REGION Network 14: Alarm and Warning
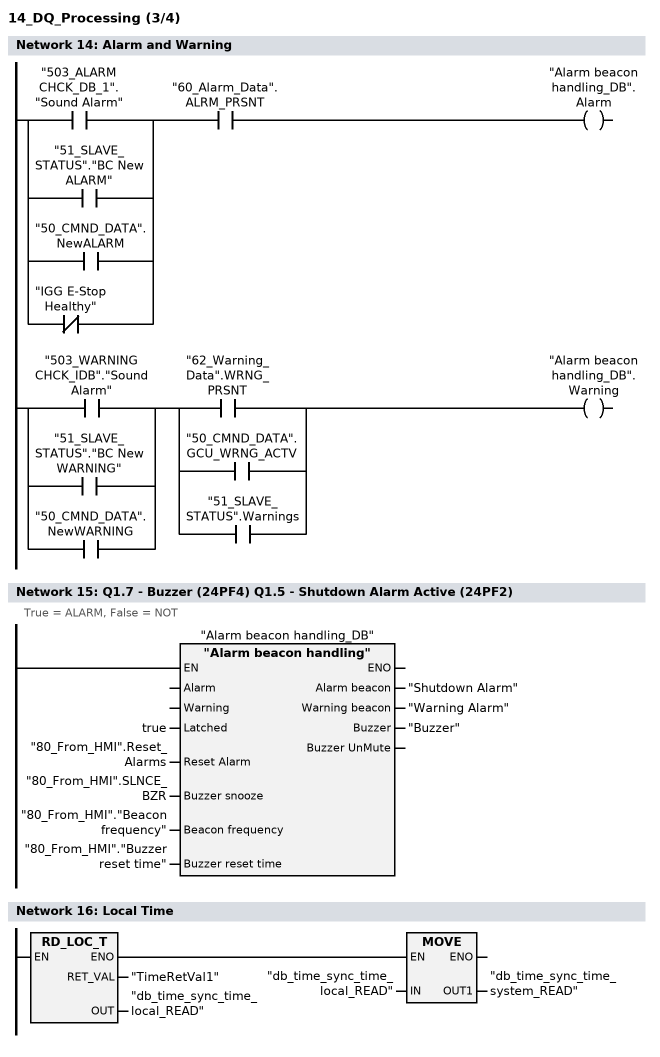
   RUNG wire#powerrail
      Contact( "503_ALARM CHCK_DB_1"."Sound Alarm" )
      wire#w1
      Contact( "60_Alarm_Data".ALRM_PRSNT )
      Coil( "Alarm beacon handling_DB".Alarm )
   END_RUNG
   RUNG wire#powerrail
      Contact( "51_SLAVE_STATUS"."BC New ALARM" )
   END_RUNG wire#w1
   RUNG wire#powerrail
      Contact( "50_CMND_DATA".NewALARM )
   END_RUNG wire#w1
   RUNG wire#powerrail
      I_Contact( "IGG E-Stop Healthy" )
   END_RUNG wire#w1
   RUNG wire#powerrail
      Contact( "503_WARNING CHCK_IDB"."Sound Alarm" )
      wire#w2
      Contact( "62_Warning_Data".WRNG_PRSNT )
      wire#w3
      Coil( "Alarm beacon handling_DB".Warning )
   END_RUNG
   RUNG wire#powerrail
      Contact( "51_SLAVE_STATUS"."BC New WARNING" )
   END_RUNG wire#w2
   RUNG wire#powerrail
      Contact( "50_CMND_DATA".NewWARNING )
   END_RUNG wire#w2
   RUNG wire#w2
      Contact( "50_CMND_DATA".GCU_WRNG_ACTV )
   END_RUNG wire#w3
   RUNG wire#w2
      Contact( "51_SLAVE_STATUS".Warnings )
   END_RUNG wire#w3
   // the same network as SCL:
   "Alarm beacon handling_DB".Alarm := ("503_ALARM CHCK_DB_1"."Sound Alarm" OR "51_SLAVE_STATUS"."BC New ALARM" OR "50_CMND_DATA".NewALARM OR NOT "IGG E-Stop Healthy") AND "60_Alarm_Data".ALRM_PRSNT;
   "Alarm beacon handling_DB".Warning := ("503_WARNING CHCK_IDB"."Sound Alarm" OR "51_SLAVE_STATUS"."BC New WARNING" OR "50_CMND_DATA".NewWARNING) AND ("62_Warning_Data".WRNG_PRSNT OR "50_CMND_DATA".GCU_WRNG_ACTV OR "51_SLAVE_STATUS".Warnings);
END_REGION

REGION Network 15: Q1.7 - Buzzer (24PF4) Q1.5 - Shutdown Alarm Active (24PF2)
   // True = ALARM, False = NOT
   RUNG wire#powerrail
      "Alarm beacon handling_DB"(Alarm :=, Warning :=, Latched := true, "Reset Alarm" := "80_From_HMI".Reset_Alarms, "Buzzer snooze" := "80_From_HMI".SLNCE_BZR, "Beacon frequency" := "80_From_HMI"."Beacon frequency", "Buzzer reset time" := "80_From_HMI"."Buzzer reset time", "Alarm beacon" => "Shutdown Alarm", "Warning beacon" => "Warning Alarm", Buzzer => "Buzzer", "Buzzer UnMute" =>)
   END_RUNG
   // the same network as SCL:
   "Alarm beacon handling_DB"(Latched := true,   // "Alarm beacon handling"
                           "Reset Alarm" := "80_From_HMI".Reset_Alarms,
                           "Buzzer snooze" := "80_From_HMI".SLNCE_BZR,
                           "Beacon frequency" := "80_From_HMI"."Beacon frequency",
                           "Buzzer reset time" := "80_From_HMI"."Buzzer reset time",
                           "Alarm beacon" => "Shutdown Alarm",
                           "Warning beacon" => "Warning Alarm",
                           Buzzer => "Buzzer");
END_REGION

REGION Network 16: Local Time
   // ENO of a box is taken as its EN; it also drops when the box reports an error
   "TimeRetVal1" := RD_LOC_T(OUT => "db_time_sync_time_local_READ");
   "db_time_sync_time_system_READ" := "db_time_sync_time_local_READ";
END_REGION

REGION Network 17: WRITE LOCAL TIME
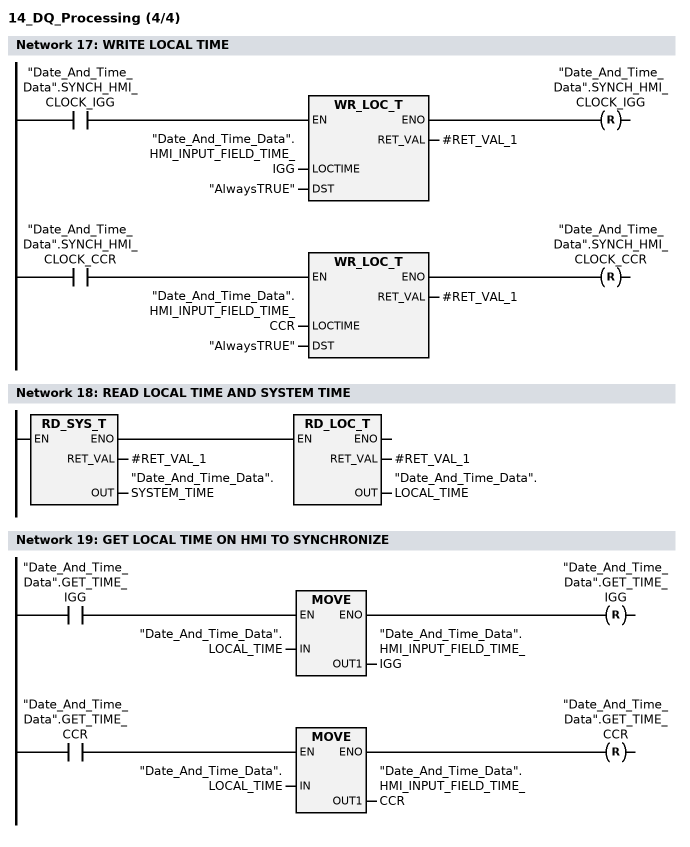
   // ENO of a box is taken as its EN; it also drops when the box reports an error
   #_w1 := "Date_And_Time_Data".SYNCH_HMI_CLOCK_IGG;
   IF #_w1 THEN
       #RET_VAL_1 := WR_LOC_T(LOCTIME := "Date_And_Time_Data".HMI_INPUT_FIELD_TIME_IGG, DST := "AlwaysTRUE");
       "Date_And_Time_Data".SYNCH_HMI_CLOCK_IGG := FALSE;
   END_IF;
   #_w2 := "Date_And_Time_Data".SYNCH_HMI_CLOCK_CCR;
   IF #_w2 THEN
       #RET_VAL_1 := WR_LOC_T(LOCTIME := "Date_And_Time_Data".HMI_INPUT_FIELD_TIME_CCR, DST := "AlwaysTRUE");
       "Date_And_Time_Data".SYNCH_HMI_CLOCK_CCR := FALSE;
   END_IF;
END_REGION

REGION Network 18: READ LOCAL TIME AND SYSTEM TIME
   // ENO of a box is taken as its EN; it also drops when the box reports an error
   #RET_VAL_1 := RD_SYS_T(OUT => "Date_And_Time_Data".SYSTEM_TIME);
   #RET_VAL_1 := RD_LOC_T(OUT => "Date_And_Time_Data".LOCAL_TIME);
END_REGION

REGION Network 19: GET LOCAL TIME ON HMI TO SYNCHRONIZE
   RUNG wire#powerrail
      Contact( "Date_And_Time_Data".GET_TIME_IGG )
      Move(in := "Date_And_Time_Data".LOCAL_TIME, out1 => "Date_And_Time_Data".HMI_INPUT_FIELD_TIME_IGG)
      R_Coil( "Date_And_Time_Data".GET_TIME_IGG )
   END_RUNG
   RUNG wire#powerrail
      Contact( "Date_And_Time_Data".GET_TIME_CCR )
      Move(in := "Date_And_Time_Data".LOCAL_TIME, out1 => "Date_And_Time_Data".HMI_INPUT_FIELD_TIME_CCR)
      R_Coil( "Date_And_Time_Data".GET_TIME_CCR )
   END_RUNG
   // the same network as SCL:
   IF "Date_And_Time_Data".GET_TIME_IGG THEN
       "Date_And_Time_Data".HMI_INPUT_FIELD_TIME_IGG := "Date_And_Time_Data".LOCAL_TIME;
       "Date_And_Time_Data".GET_TIME_IGG := FALSE;
   END_IF;
   IF "Date_And_Time_Data".GET_TIME_CCR THEN
       "Date_And_Time_Data".HMI_INPUT_FIELD_TIME_CCR := "Date_And_Time_Data".LOCAL_TIME;
       "Date_And_Time_Data".GET_TIME_CCR := FALSE;
   END_IF;
END_REGION
END_FUNCTION

FUNCTION "16_AQ_Processing" : Void   // FC16, LAD
TITLE = Analogue Output Processing
{ S7_Optimized_Access := 'TRUE' }
AUTHOR : JRS
VERSION : 0.1
// To process code outputs prior to physical connection
BEGIN

REGION Network 1: QW98 - Vent Valve Position Control (CV-403)
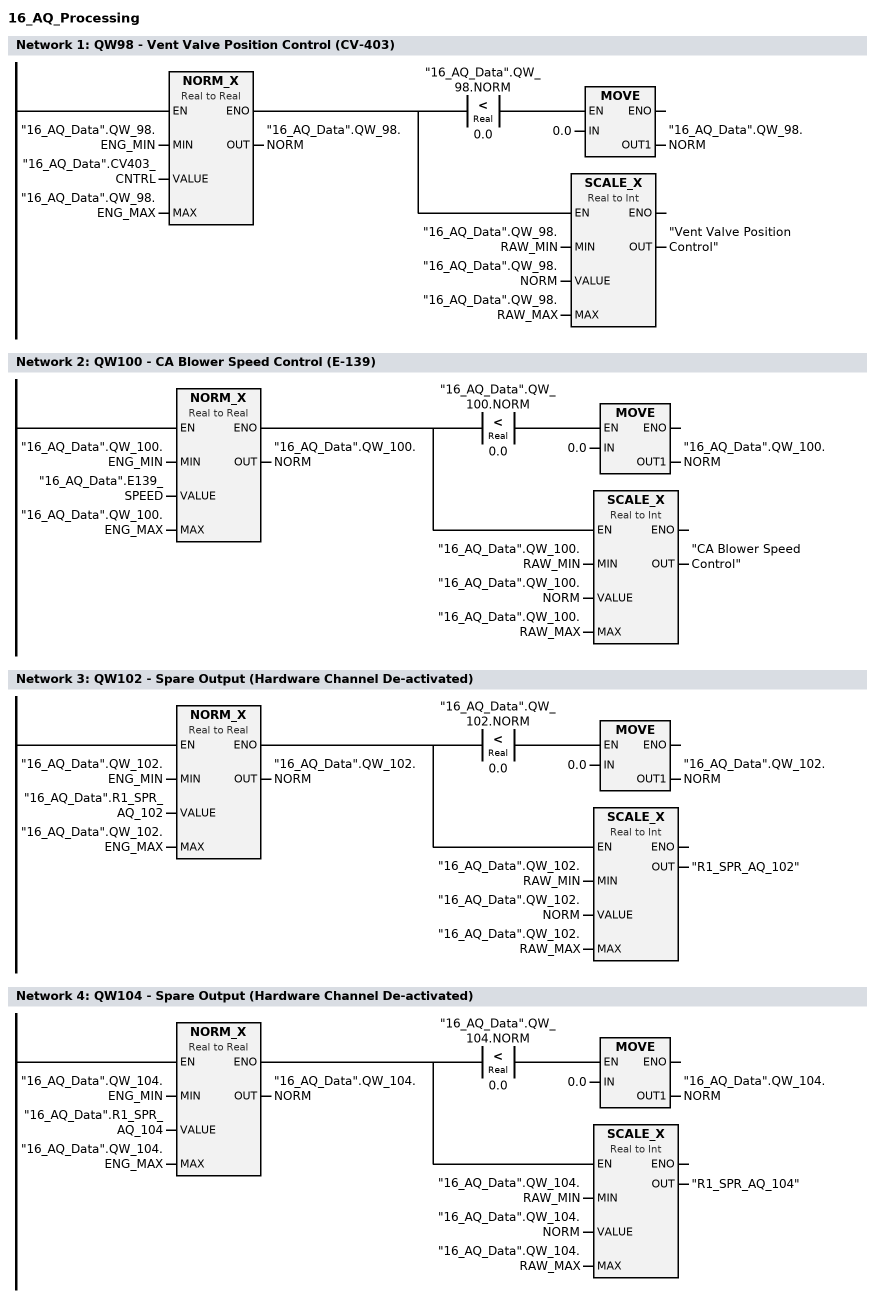
   RUNG wire#powerrail
      { S7_Templates := "[SrcType := Real, DestType := Real]" } Normalize(min := "16_AQ_Data".QW_98.ENG_MIN, value := "16_AQ_Data".CV403_CNTRL, max := "16_AQ_Data".QW_98.ENG_MAX, out => "16_AQ_Data".QW_98.NORM)
      wire#w1
      { S7_Templates := "SrcType := Real" } LT_Contact(in1 := "16_AQ_Data".QW_98.NORM, in2 := 0.0)
      Move(in := 0.0, out1 => "16_AQ_Data".QW_98.NORM)
   END_RUNG
   RUNG wire#w1
      { S7_Templates := "[SrcType := Real, DestType := Int]" } Scale(min := "16_AQ_Data".QW_98.RAW_MIN, value := "16_AQ_Data".QW_98.NORM, max := "16_AQ_Data".QW_98.RAW_MAX, out => "Vent Valve Position Control")
   END_RUNG
   // the same network as SCL:
   "16_AQ_Data".QW_98.NORM := NORM_X(MIN := "16_AQ_Data".QW_98.ENG_MIN, VALUE := "16_AQ_Data".CV403_CNTRL, MAX := "16_AQ_Data".QW_98.ENG_MAX);
   IF "16_AQ_Data".QW_98.NORM < 0.0 THEN "16_AQ_Data".QW_98.NORM := 0.0; END_IF;
   "Vent Valve Position Control" := SCALE_X(MIN := "16_AQ_Data".QW_98.RAW_MIN, VALUE := "16_AQ_Data".QW_98.NORM, MAX := "16_AQ_Data".QW_98.RAW_MAX);
END_REGION

REGION Network 2: QW100 - CA Blower Speed Control (E-139)
   RUNG wire#powerrail
      { S7_Templates := "[SrcType := Real, DestType := Real]" } Normalize(min := "16_AQ_Data".QW_100.ENG_MIN, value := "16_AQ_Data".E139_SPEED, max := "16_AQ_Data".QW_100.ENG_MAX, out => "16_AQ_Data".QW_100.NORM)
      wire#w1
      { S7_Templates := "SrcType := Real" } LT_Contact(in1 := "16_AQ_Data".QW_100.NORM, in2 := 0.0)
      Move(in := 0.0, out1 => "16_AQ_Data".QW_100.NORM)
   END_RUNG
   RUNG wire#w1
      { S7_Templates := "[SrcType := Real, DestType := Int]" } Scale(min := "16_AQ_Data".QW_100.RAW_MIN, value := "16_AQ_Data".QW_100.NORM, max := "16_AQ_Data".QW_100.RAW_MAX, out => "CA Blower Speed Control")
   END_RUNG
   // the same network as SCL:
   "16_AQ_Data".QW_100.NORM := NORM_X(MIN := "16_AQ_Data".QW_100.ENG_MIN, VALUE := "16_AQ_Data".E139_SPEED, MAX := "16_AQ_Data".QW_100.ENG_MAX);
   IF "16_AQ_Data".QW_100.NORM < 0.0 THEN "16_AQ_Data".QW_100.NORM := 0.0; END_IF;
   "CA Blower Speed Control" := SCALE_X(MIN := "16_AQ_Data".QW_100.RAW_MIN, VALUE := "16_AQ_Data".QW_100.NORM, MAX := "16_AQ_Data".QW_100.RAW_MAX);
END_REGION

REGION Network 3: QW102 - Spare Output (Hardware Channel De-activated)
   RUNG wire#powerrail
      { S7_Templates := "[SrcType := Real, DestType := Real]" } Normalize(min := "16_AQ_Data".QW_102.ENG_MIN, value := "16_AQ_Data".R1_SPR_AQ_102, max := "16_AQ_Data".QW_102.ENG_MAX, out => "16_AQ_Data".QW_102.NORM)
      wire#w1
      { S7_Templates := "SrcType := Real" } LT_Contact(in1 := "16_AQ_Data".QW_102.NORM, in2 := 0.0)
      Move(in := 0.0, out1 => "16_AQ_Data".QW_102.NORM)
   END_RUNG
   RUNG wire#w1
      { S7_Templates := "[SrcType := Real, DestType := Int]" } Scale(min := "16_AQ_Data".QW_102.RAW_MIN, value := "16_AQ_Data".QW_102.NORM, max := "16_AQ_Data".QW_102.RAW_MAX, out => "R1_SPR_AQ_102")
   END_RUNG
   // the same network as SCL:
   "16_AQ_Data".QW_102.NORM := NORM_X(MIN := "16_AQ_Data".QW_102.ENG_MIN, VALUE := "16_AQ_Data".R1_SPR_AQ_102, MAX := "16_AQ_Data".QW_102.ENG_MAX);
   IF "16_AQ_Data".QW_102.NORM < 0.0 THEN "16_AQ_Data".QW_102.NORM := 0.0; END_IF;
   "R1_SPR_AQ_102" := SCALE_X(MIN := "16_AQ_Data".QW_102.RAW_MIN, VALUE := "16_AQ_Data".QW_102.NORM, MAX := "16_AQ_Data".QW_102.RAW_MAX);
END_REGION

REGION Network 4: QW104 - Spare Output (Hardware Channel De-activated)
   RUNG wire#powerrail
      { S7_Templates := "[SrcType := Real, DestType := Real]" } Normalize(min := "16_AQ_Data".QW_104.ENG_MIN, value := "16_AQ_Data".R1_SPR_AQ_104, max := "16_AQ_Data".QW_104.ENG_MAX, out => "16_AQ_Data".QW_104.NORM)
      wire#w1
      { S7_Templates := "SrcType := Real" } LT_Contact(in1 := "16_AQ_Data".QW_104.NORM, in2 := 0.0)
      Move(in := 0.0, out1 => "16_AQ_Data".QW_104.NORM)
   END_RUNG
   RUNG wire#w1
      { S7_Templates := "[SrcType := Real, DestType := Int]" } Scale(min := "16_AQ_Data".QW_104.RAW_MIN, value := "16_AQ_Data".QW_104.NORM, max := "16_AQ_Data".QW_104.RAW_MAX, out => "R1_SPR_AQ_104")
   END_RUNG
   // the same network as SCL:
   "16_AQ_Data".QW_104.NORM := NORM_X(MIN := "16_AQ_Data".QW_104.ENG_MIN, VALUE := "16_AQ_Data".R1_SPR_AQ_104, MAX := "16_AQ_Data".QW_104.ENG_MAX);
   IF "16_AQ_Data".QW_104.NORM < 0.0 THEN "16_AQ_Data".QW_104.NORM := 0.0; END_IF;
   "R1_SPR_AQ_104" := SCALE_X(MIN := "16_AQ_Data".QW_104.RAW_MIN, VALUE := "16_AQ_Data".QW_104.NORM, MAX := "16_AQ_Data".QW_104.RAW_MAX);
END_REGION
END_FUNCTION

FUNCTION "19_AUTO_CMNDS" : Void   // FC19, LAD
TITLE = Automatic Output Commands
{ S7_Optimized_Access := 'TRUE' }
AUTHOR : JRS
VERSION : 0.1
// To process automatic output commands prior to output processing
   VAR_TEMP   // added for the SCL form of the ladder/FBD networks
      _w1 : Bool;
      _w2 : Bool;
   END_VAR
BEGIN

REGION Network 1: Fuel Pumps Control
   // Demand from sequence     ...changed from 80 to 140
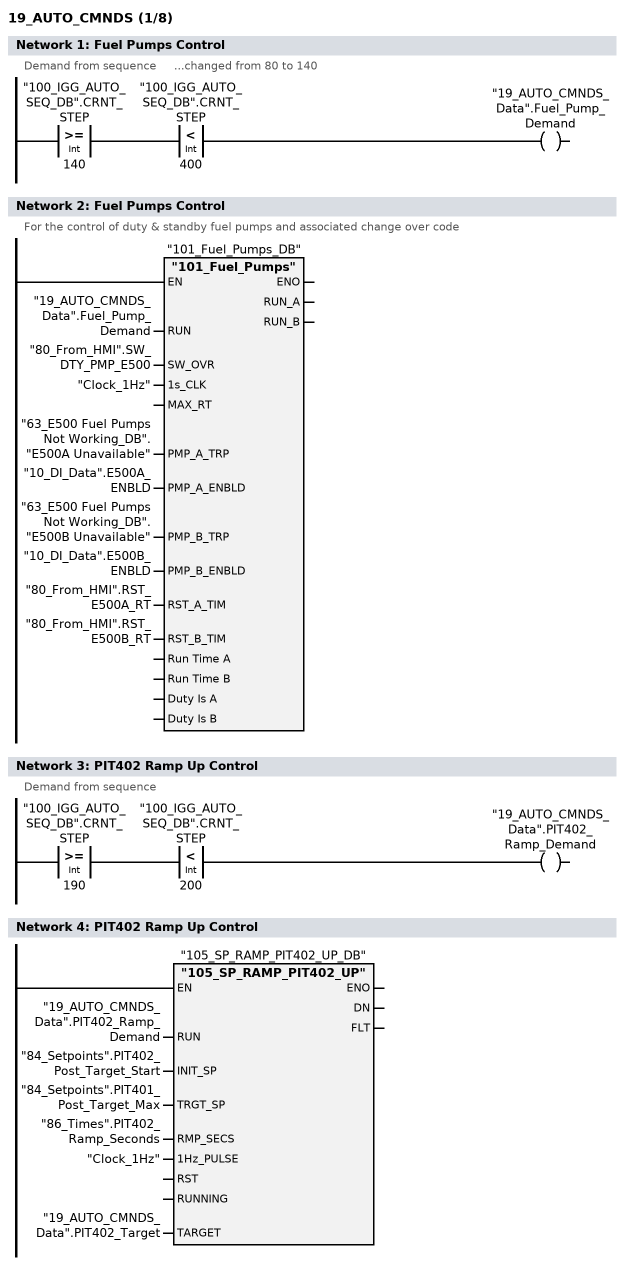
   RUNG wire#powerrail
      { S7_Templates := "SrcType := Int" } GE_Contact(in1 := "100_IGG_AUTO_SEQ_DB".CRNT_STEP, in2 := 140)
      { S7_Templates := "SrcType := Int" } LT_Contact(in1 := "100_IGG_AUTO_SEQ_DB".CRNT_STEP, in2 := 400)
      Coil( "19_AUTO_CMNDS_Data".Fuel_Pump_Demand )
   END_RUNG
   // the same network as SCL:
   "19_AUTO_CMNDS_Data".Fuel_Pump_Demand := ("100_IGG_AUTO_SEQ_DB".CRNT_STEP >= 140) AND ("100_IGG_AUTO_SEQ_DB".CRNT_STEP < 400);
END_REGION

REGION Network 2: Fuel Pumps Control
   // For the control of duty & standby fuel pumps and associated change over code
   RUNG wire#powerrail
      "101_Fuel_Pumps_DB"(RUN := "19_AUTO_CMNDS_Data".Fuel_Pump_Demand, SW_OVR := "80_From_HMI".SW_DTY_PMP_E500, "1s_CLK" := "Clock_1Hz", MAX_RT :=, PMP_A_TRP := "63_E500 Fuel Pumps Not Working_DB"."E500A Unavailable", PMP_A_ENBLD := "10_DI_Data".E500A_ENBLD, PMP_B_TRP := "63_E500 Fuel Pumps Not Working_DB"."E500B Unavailable", PMP_B_ENBLD := "10_DI_Data".E500B_ENBLD, RST_A_TIM := "80_From_HMI".RST_E500A_RT, RST_B_TIM := "80_From_HMI".RST_E500B_RT, "Run Time A" :=, "Run Time B" :=, "Duty Is A" :=, "Duty Is B" :=, RUN_A =>, RUN_B =>)
   END_RUNG
   // the same network as SCL:
   "101_Fuel_Pumps_DB"(RUN := "19_AUTO_CMNDS_Data".Fuel_Pump_Demand,   // "101_Fuel_Pumps"
                       SW_OVR := "80_From_HMI".SW_DTY_PMP_E500,
                       "1s_CLK" := "Clock_1Hz",
                       PMP_A_TRP := "63_E500 Fuel Pumps Not Working_DB"."E500A Unavailable",
                       PMP_A_ENBLD := "10_DI_Data".E500A_ENBLD,
                       PMP_B_TRP := "63_E500 Fuel Pumps Not Working_DB"."E500B Unavailable",
                       PMP_B_ENBLD := "10_DI_Data".E500B_ENBLD,
                       RST_A_TIM := "80_From_HMI".RST_E500A_RT,
                       RST_B_TIM := "80_From_HMI".RST_E500B_RT);
END_REGION

REGION Network 3: PIT402 Ramp Up Control
   // Demand from sequence
   RUNG wire#powerrail
      { S7_Templates := "SrcType := Int" } GE_Contact(in1 := "100_IGG_AUTO_SEQ_DB".CRNT_STEP, in2 := 190)
      { S7_Templates := "SrcType := Int" } LT_Contact(in1 := "100_IGG_AUTO_SEQ_DB".CRNT_STEP, in2 := 200)
      Coil( "19_AUTO_CMNDS_Data".PIT402_Ramp_Demand )
   END_RUNG
   // the same network as SCL:
   "19_AUTO_CMNDS_Data".PIT402_Ramp_Demand := ("100_IGG_AUTO_SEQ_DB".CRNT_STEP >= 190) AND ("100_IGG_AUTO_SEQ_DB".CRNT_STEP < 200);
END_REGION

REGION Network 4: PIT402 Ramp Up Control
   RUNG wire#powerrail
      "105_SP_RAMP_PIT402_UP_DB"(RUN := "19_AUTO_CMNDS_Data".PIT402_Ramp_Demand, INIT_SP := "84_Setpoints".PIT402_Post_Target_Start, TRGT_SP := "84_Setpoints".PIT401_Post_Target_Max, RMP_SECS := "86_Times".PIT402_Ramp_Seconds, "1Hz_PULSE" := "Clock_1Hz", RST :=, RUNNING :=, TARGET := "19_AUTO_CMNDS_Data".PIT402_Target, DN =>, FLT =>)
   END_RUNG
   // the same network as SCL:
   "105_SP_RAMP_PIT402_UP_DB"(RUN := "19_AUTO_CMNDS_Data".PIT402_Ramp_Demand,   // "105_SP_RAMP_PIT402_UP"
                           INIT_SP := "84_Setpoints".PIT402_Post_Target_Start,
                           TRGT_SP := "84_Setpoints".PIT401_Post_Target_Max,
                           RMP_SECS := "86_Times".PIT402_Ramp_Seconds,
                           "1Hz_PULSE" := "Clock_1Hz",
                           TARGET := "19_AUTO_CMNDS_Data".PIT402_Target);
END_REGION

REGION Network 5: PIT402 Ramp Down Control
   // Demand from sequence
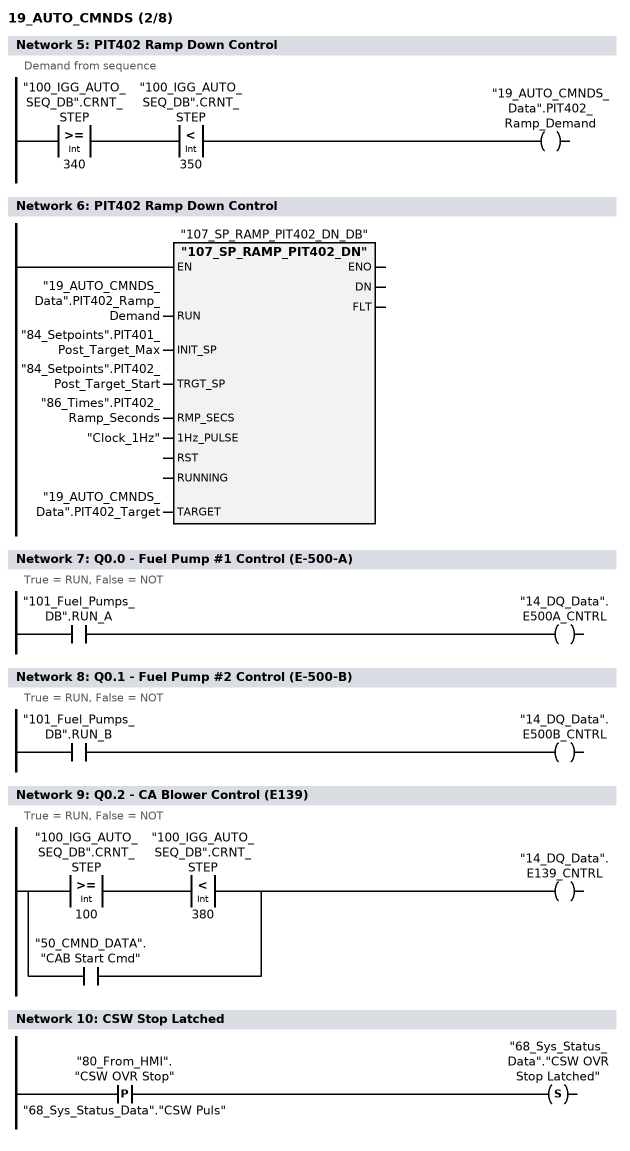
   RUNG wire#powerrail
      { S7_Templates := "SrcType := Int" } GE_Contact(in1 := "100_IGG_AUTO_SEQ_DB".CRNT_STEP, in2 := 340)
      { S7_Templates := "SrcType := Int" } LT_Contact(in1 := "100_IGG_AUTO_SEQ_DB".CRNT_STEP, in2 := 350)
      Coil( "19_AUTO_CMNDS_Data".PIT402_Ramp_Demand )
   END_RUNG
   // the same network as SCL:
   "19_AUTO_CMNDS_Data".PIT402_Ramp_Demand := ("100_IGG_AUTO_SEQ_DB".CRNT_STEP >= 340) AND ("100_IGG_AUTO_SEQ_DB".CRNT_STEP < 350);
END_REGION

REGION Network 6: PIT402 Ramp Down Control
   RUNG wire#powerrail
      "107_SP_RAMP_PIT402_DN_DB"(RUN := "19_AUTO_CMNDS_Data".PIT402_Ramp_Demand, INIT_SP := "84_Setpoints".PIT401_Post_Target_Max, TRGT_SP := "84_Setpoints".PIT402_Post_Target_Start, RMP_SECS := "86_Times".PIT402_Ramp_Seconds, "1Hz_PULSE" := "Clock_1Hz", RST :=, RUNNING :=, TARGET := "19_AUTO_CMNDS_Data".PIT402_Target, DN =>, FLT =>)
   END_RUNG
   // the same network as SCL:
   "107_SP_RAMP_PIT402_DN_DB"(RUN := "19_AUTO_CMNDS_Data".PIT402_Ramp_Demand,   // "107_SP_RAMP_PIT402_DN"
                           INIT_SP := "84_Setpoints".PIT401_Post_Target_Max,
                           TRGT_SP := "84_Setpoints".PIT402_Post_Target_Start,
                           RMP_SECS := "86_Times".PIT402_Ramp_Seconds,
                           "1Hz_PULSE" := "Clock_1Hz",
                           TARGET := "19_AUTO_CMNDS_Data".PIT402_Target);
END_REGION

REGION Network 7: Q0.0 - Fuel Pump #1 Control (E-500-A)
   // True = RUN, False = NOT
   RUNG wire#powerrail
      Contact( "101_Fuel_Pumps_DB".RUN_A )
      Coil( "14_DQ_Data".E500A_CNTRL )
   END_RUNG
   // the same network as SCL:
   "14_DQ_Data".E500A_CNTRL := "101_Fuel_Pumps_DB".RUN_A;
END_REGION

REGION Network 8: Q0.1 - Fuel Pump #2 Control (E-500-B)
   // True = RUN, False = NOT
   RUNG wire#powerrail
      Contact( "101_Fuel_Pumps_DB".RUN_B )
      Coil( "14_DQ_Data".E500B_CNTRL )
   END_RUNG
   // the same network as SCL:
   "14_DQ_Data".E500B_CNTRL := "101_Fuel_Pumps_DB".RUN_B;
END_REGION

REGION Network 9: Q0.2 - CA Blower Control (E139)
   // True = RUN, False = NOT
   RUNG wire#powerrail
      { S7_Templates := "SrcType := Int" } GE_Contact(in1 := "100_IGG_AUTO_SEQ_DB".CRNT_STEP, in2 := 100)
      { S7_Templates := "SrcType := Int" } LT_Contact(in1 := "100_IGG_AUTO_SEQ_DB".CRNT_STEP, in2 := 380)
      wire#w1
      Coil( "14_DQ_Data".E139_CNTRL )
   END_RUNG
   RUNG wire#powerrail
      Contact( "50_CMND_DATA"."CAB Start Cmd" )
   END_RUNG wire#w1
   // the same network as SCL:
   "14_DQ_Data".E139_CNTRL := (("100_IGG_AUTO_SEQ_DB".CRNT_STEP >= 100) AND ("100_IGG_AUTO_SEQ_DB".CRNT_STEP < 380)) OR "50_CMND_DATA"."CAB Start Cmd";
END_REGION

REGION Network 10: CSW Stop Latched
   RUNG wire#powerrail
      P_Contact(operand := "80_From_HMI"."CSW OVR Stop", bit := "68_Sys_Status_Data"."CSW Puls")
      S_Coil( "68_Sys_Status_Data"."CSW OVR Stop Latched" )
   END_RUNG
   // the same network as SCL:
   #_w1 := "80_From_HMI"."CSW OVR Stop" AND NOT "68_Sys_Status_Data"."CSW Puls";   // rising edge of "80_From_HMI"."CSW OVR Stop"
   "68_Sys_Status_Data"."CSW Puls" := "80_From_HMI"."CSW OVR Stop";
   IF #_w1 THEN "68_Sys_Status_Data"."CSW OVR Stop Latched" := TRUE; END_IF;
END_REGION

REGION Network 11: Q0.3 - Cooling Sea Water (CSW) Inlet Valves Control (CV311)
   // True = OPEN, False = CLOSE
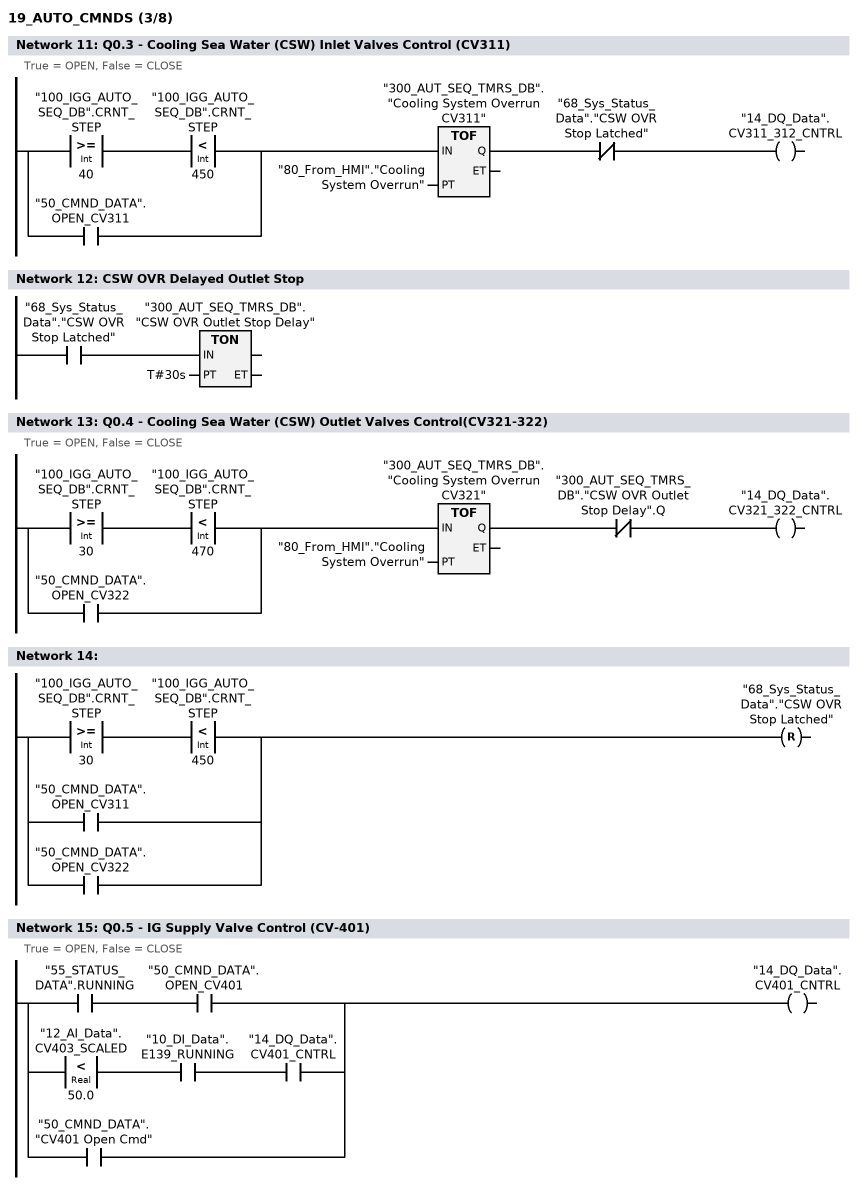
   "300_AUT_SEQ_TMRS_DB"."Cooling System Overrun CV311".TOF(IN := (("100_IGG_AUTO_SEQ_DB".CRNT_STEP >= 40) AND ("100_IGG_AUTO_SEQ_DB".CRNT_STEP < 450)) OR "50_CMND_DATA".OPEN_CV311,
                           PT := "80_From_HMI"."Cooling System Overrun");
   "14_DQ_Data".CV311_312_CNTRL := "300_AUT_SEQ_TMRS_DB"."Cooling System Overrun CV311".Q AND NOT "68_Sys_Status_Data"."CSW OVR Stop Latched";
END_REGION

REGION Network 12: CSW OVR Delayed Outlet Stop
   "300_AUT_SEQ_TMRS_DB"."CSW OVR Outlet Stop Delay".TON(IN := "68_Sys_Status_Data"."CSW OVR Stop Latched",
                           PT := T#30s);
END_REGION

REGION Network 13: Q0.4 - Cooling Sea Water (CSW) Outlet Valves Control(CV321-322)
   // True = OPEN, False = CLOSE
   "300_AUT_SEQ_TMRS_DB"."Cooling System Overrun CV321".TOF(IN := (("100_IGG_AUTO_SEQ_DB".CRNT_STEP >= 30) AND ("100_IGG_AUTO_SEQ_DB".CRNT_STEP < 470)) OR "50_CMND_DATA".OPEN_CV322,
                           PT := "80_From_HMI"."Cooling System Overrun");
   "14_DQ_Data".CV321_322_CNTRL := "300_AUT_SEQ_TMRS_DB"."Cooling System Overrun CV321".Q AND NOT "300_AUT_SEQ_TMRS_DB"."CSW OVR Outlet Stop Delay".Q;
END_REGION

REGION Network 14
   RUNG wire#powerrail
      { S7_Templates := "SrcType := Int" } GE_Contact(in1 := "100_IGG_AUTO_SEQ_DB".CRNT_STEP, in2 := 30)
      { S7_Templates := "SrcType := Int" } LT_Contact(in1 := "100_IGG_AUTO_SEQ_DB".CRNT_STEP, in2 := 450)
      wire#w1
      R_Coil( "68_Sys_Status_Data"."CSW OVR Stop Latched" )
   END_RUNG
   RUNG wire#powerrail
      Contact( "50_CMND_DATA".OPEN_CV311 )
   END_RUNG wire#w1
   RUNG wire#powerrail
      Contact( "50_CMND_DATA".OPEN_CV322 )
   END_RUNG wire#w1
   // the same network as SCL:
   IF (("100_IGG_AUTO_SEQ_DB".CRNT_STEP >= 30) AND ("100_IGG_AUTO_SEQ_DB".CRNT_STEP < 450)) OR "50_CMND_DATA".OPEN_CV311 OR "50_CMND_DATA".OPEN_CV322 THEN
       "68_Sys_Status_Data"."CSW OVR Stop Latched" := FALSE;
   END_IF;
END_REGION

REGION Network 15: Q0.5 - IG Supply Valve Control (CV-401)
   // True = OPEN, False = CLOSE
   RUNG wire#powerrail
      Contact( "55_STATUS_DATA".RUNNING )
      Contact( "50_CMND_DATA".OPEN_CV401 )
      wire#w1
      Coil( "14_DQ_Data".CV401_CNTRL )
   END_RUNG
   RUNG wire#powerrail
      { S7_Templates := "SrcType := Real" } LT_Contact(in1 := "12_AI_Data".CV403_SCALED, in2 := 50.0)
      Contact( "10_DI_Data".E139_RUNNING )
      Contact( "14_DQ_Data".CV401_CNTRL )
   END_RUNG wire#w1
   RUNG wire#powerrail
      Contact( "50_CMND_DATA"."CV401 Open Cmd" )
   END_RUNG wire#w1
   // the same network as SCL:
   "14_DQ_Data".CV401_CNTRL := ("55_STATUS_DATA".RUNNING AND "50_CMND_DATA".OPEN_CV401) OR (("12_AI_Data".CV403_SCALED < 50.0) AND "10_DI_Data".E139_RUNNING AND "14_DQ_Data".CV401_CNTRL) OR "50_CMND_DATA"."CV401 Open Cmd";
END_REGION

REGION Network 16: Q0.6 - Cargo Blanketing/BWTS Valve Control (CV431/432)
   // True = RUN, False = NOT
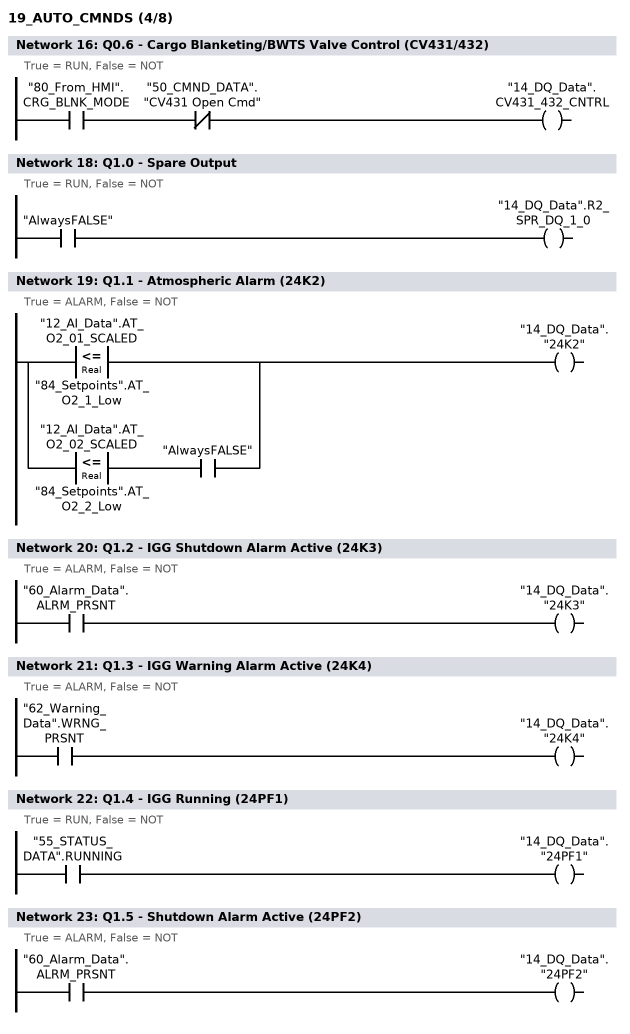
   RUNG wire#powerrail
      Contact( "80_From_HMI".CRG_BLNK_MODE )
      I_Contact( "50_CMND_DATA"."CV431 Open Cmd" )
      Coil( "14_DQ_Data".CV431_432_CNTRL )
   END_RUNG
   // the same network as SCL:
   "14_DQ_Data".CV431_432_CNTRL := "80_From_HMI".CRG_BLNK_MODE AND NOT "50_CMND_DATA"."CV431 Open Cmd";
END_REGION

REGION Network 17: Q0.7
   // True = RUN, False = NOT
END_REGION

REGION Network 18: Q1.0 - Spare Output
   // True = RUN, False = NOT
   RUNG wire#powerrail
      Contact( "AlwaysFALSE" )
      Coil( "14_DQ_Data".R2_SPR_DQ_1_0 )
   END_RUNG
   // the same network as SCL:
   "14_DQ_Data".R2_SPR_DQ_1_0 := "AlwaysFALSE";
END_REGION

REGION Network 19: Q1.1 - Atmospheric Alarm (24K2)
   // True = ALARM, False = NOT
   RUNG wire#powerrail
      { S7_Templates := "SrcType := Real" } LE_Contact(in1 := "12_AI_Data".AT_O2_01_SCALED, in2 := "84_Setpoints".AT_O2_1_Low)
      wire#w1
      Coil( "14_DQ_Data"."24K2" )
   END_RUNG
   RUNG wire#powerrail
      { S7_Templates := "SrcType := Real" } LE_Contact(in1 := "12_AI_Data".AT_O2_02_SCALED, in2 := "84_Setpoints".AT_O2_2_Low)
      Contact( "AlwaysFALSE" )
   END_RUNG wire#w1
   // the same network as SCL:
   "14_DQ_Data"."24K2" := ("12_AI_Data".AT_O2_01_SCALED <= "84_Setpoints".AT_O2_1_Low) OR (("12_AI_Data".AT_O2_02_SCALED <= "84_Setpoints".AT_O2_2_Low) AND "AlwaysFALSE");
END_REGION

REGION Network 20: Q1.2 - IGG Shutdown Alarm Active (24K3)
   // True = ALARM, False = NOT
   RUNG wire#powerrail
      Contact( "60_Alarm_Data".ALRM_PRSNT )
      Coil( "14_DQ_Data"."24K3" )
   END_RUNG
   // the same network as SCL:
   "14_DQ_Data"."24K3" := "60_Alarm_Data".ALRM_PRSNT;
END_REGION

REGION Network 21: Q1.3 - IGG Warning Alarm Active (24K4)
   // True = ALARM, False = NOT
   RUNG wire#powerrail
      Contact( "62_Warning_Data".WRNG_PRSNT )
      Coil( "14_DQ_Data"."24K4" )
   END_RUNG
   // the same network as SCL:
   "14_DQ_Data"."24K4" := "62_Warning_Data".WRNG_PRSNT;
END_REGION

REGION Network 22: Q1.4 - IGG Running (24PF1)
   // True = RUN, False = NOT
   RUNG wire#powerrail
      Contact( "55_STATUS_DATA".RUNNING )
      Coil( "14_DQ_Data"."24PF1" )
   END_RUNG
   // the same network as SCL:
   "14_DQ_Data"."24PF1" := "55_STATUS_DATA".RUNNING;
END_REGION

REGION Network 23: Q1.5 - Shutdown Alarm Active (24PF2)
   // True = ALARM, False = NOT
   RUNG wire#powerrail
      Contact( "60_Alarm_Data".ALRM_PRSNT )
      Coil( "14_DQ_Data"."24PF2" )
   END_RUNG
   // the same network as SCL:
   "14_DQ_Data"."24PF2" := "60_Alarm_Data".ALRM_PRSNT;
END_REGION

REGION Network 24: Q1.6 - Warning Alarm Active (24PF3)
   // True = ALARM, False = NOT
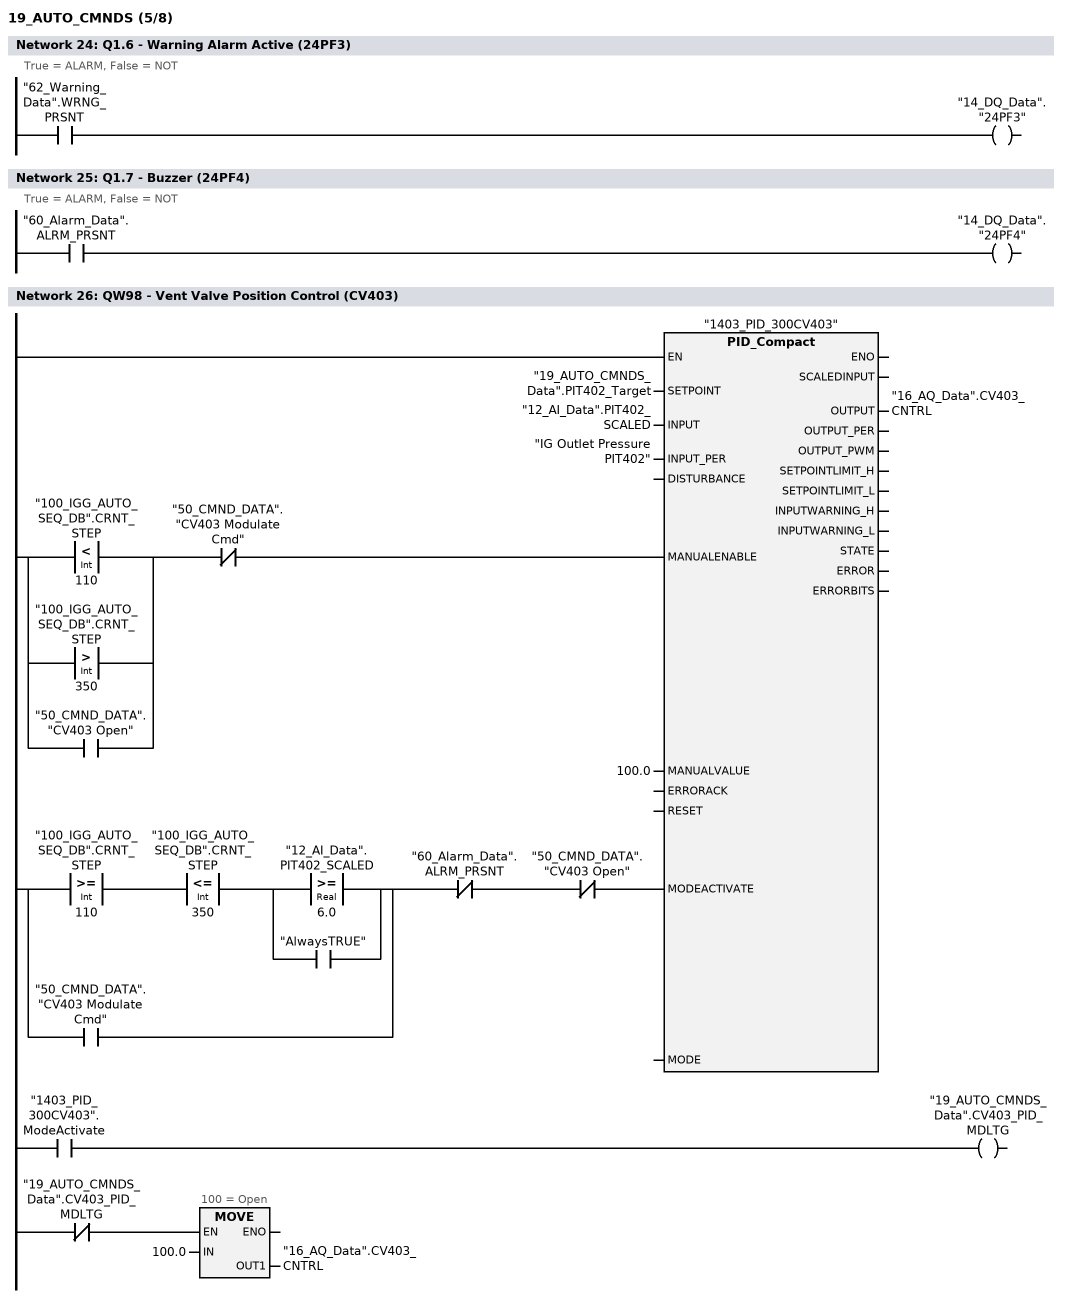
   RUNG wire#powerrail
      Contact( "62_Warning_Data".WRNG_PRSNT )
      Coil( "14_DQ_Data"."24PF3" )
   END_RUNG
   // the same network as SCL:
   "14_DQ_Data"."24PF3" := "62_Warning_Data".WRNG_PRSNT;
END_REGION

REGION Network 25: Q1.7 - Buzzer (24PF4)
   // True = ALARM, False = NOT
   RUNG wire#powerrail
      Contact( "60_Alarm_Data".ALRM_PRSNT )
      Coil( "14_DQ_Data"."24PF4" )
   END_RUNG
   // the same network as SCL:
   "14_DQ_Data"."24PF4" := "60_Alarm_Data".ALRM_PRSNT;
END_REGION

REGION Network 26: QW98 - Vent Valve Position Control (CV403)
   "1403_PID_300CV403"(Setpoint := "19_AUTO_CMNDS_Data".PIT402_Target,   // PID_Compact
                       Input := "12_AI_Data".PIT402_SCALED,
                       Input_PER := "IG Outlet Pressure PIT402",
                       ManualEnable := (("100_IGG_AUTO_SEQ_DB".CRNT_STEP < 110) OR ("100_IGG_AUTO_SEQ_DB".CRNT_STEP > 350) OR "50_CMND_DATA"."CV403 Open") AND NOT "50_CMND_DATA"."CV403 Modulate Cmd",
                       ManualValue := 100.0,
                       ModeActivate := ((("100_IGG_AUTO_SEQ_DB".CRNT_STEP >= 110) AND ("100_IGG_AUTO_SEQ_DB".CRNT_STEP <= 350) AND (("12_AI_Data".PIT402_SCALED >= 6.0) OR "AlwaysTRUE")) OR "50_CMND_DATA"."CV403 Modulate Cmd") AND NOT "60_Alarm_Data".ALRM_PRSNT AND NOT "50_CMND_DATA"."CV403 Open",
                       Output => "16_AQ_Data".CV403_CNTRL);
   "19_AUTO_CMNDS_Data".CV403_PID_MDLTG := "1403_PID_300CV403".ModeActivate;
   IF NOT "19_AUTO_CMNDS_Data".CV403_PID_MDLTG THEN
       "16_AQ_Data".CV403_CNTRL := 100.0;   // 100 = Open
   END_IF;
END_REGION

REGION Network 27: QW100 - CA Blower Speed Control (E-139)